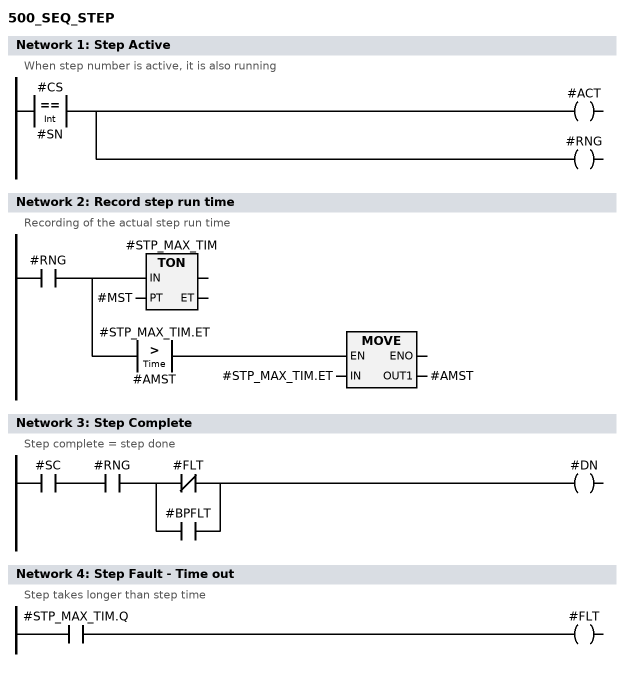
   RUNG wire#powerrail
      { S7_Templates := "SrcType := Int" } EQ_Contact(in1 := #CS, in2 := #SN)
      wire#w1
      Coil( #ACT )
   END_RUNG
   RUNG wire#w1
      Coil( #RNG )
   END_RUNG
   // the same network as SCL:
   #ACT := #CS = #SN;
   #RNG := #ACT;
END_REGION

REGION Network 2: Record step run time
   // Recording of the actual step run time
   #STP_MAX_TIM(IN := #RNG, PT := #MST);   // TON
   IF #RNG AND (#STP_MAX_TIM.ET > #AMST) THEN #AMST := #STP_MAX_TIM.ET; END_IF;
END_REGION

REGION Network 3: Step Complete
   // Step complete = step done
   RUNG wire#powerrail
      Contact( #SC )
      Contact( #RNG )
      wire#w1
      I_Contact( #FLT )
      wire#w2
      Coil( #DN )
   END_RUNG
   RUNG wire#w1
      Contact( #BPFLT )
   END_RUNG wire#w2
   // the same network as SCL:
   #DN := #SC AND #RNG AND (NOT #FLT OR #BPFLT);
END_REGION

REGION Network 4: Step Fault - Time out
   // Step takes longer than step time
   RUNG wire#powerrail
      Contact( #STP_MAX_TIM.Q )
      Coil( #FLT )
   END_RUNG
   // the same network as SCL:
   #FLT := #STP_MAX_TIM.Q;
END_REGION
END_FUNCTION_BLOCK

FUNCTION_BLOCK "501_VLV_CHK"   // FB501, LAD
TITLE = Valve Check
{ S7_Optimized_Access := 'TRUE' }
AUTHOR : JRS
VERSION : 0.1
// To check for the correct operation of a vlave
   VAR_INPUT
      DMND : Bool;   // Demand
      NO_TYPE : Bool;   // Valve type = open without demand
      NC_TYPE : Bool;   // Valve type = closed without demand
      MAX_MOV_TIM : Time := T#1s;   // Maximum movement time
      OPN_SNSR : Bool;   // Valve open confirmed
      CLS_SNSR : Bool;   // Valve closed confirmed
   END_VAR
   VAR_OUTPUT
      HELTHY : Bool;   // Valve is healthy
      FAULT : Bool;   // Valve is faulty
      CNFG_ERR : Bool;   // Configuration error
   END_VAR
   VAR
      IDLE_FLT : Bool;   // No demand fault
      DMND_FLT : Bool;   // Demand fault
      TRVL_TIME_FLT : Bool;   // Both sensors missing
      SNSR_FLT : Bool;   // Sensor conflicts
      TRVL_TIME : TON_TIME;   // Travel timer
   END_VAR
   // TRVL_TIME.PT := T#1s;
BEGIN

REGION Network 1: Idle Fault
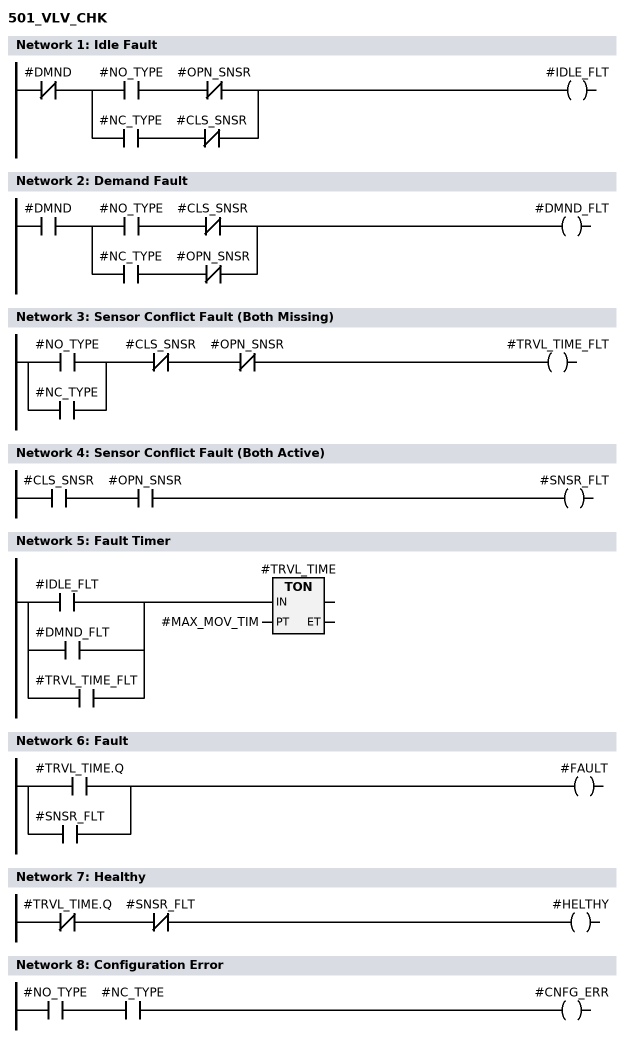
   RUNG wire#powerrail
      I_Contact( #DMND )
      wire#w1
      Contact( #NO_TYPE )
      I_Contact( #OPN_SNSR )
      wire#w2
      Coil( #IDLE_FLT )
   END_RUNG
   RUNG wire#w1
      Contact( #NC_TYPE )
      I_Contact( #CLS_SNSR )
   END_RUNG wire#w2
   // the same network as SCL:
   #IDLE_FLT := NOT #DMND AND ((#NO_TYPE AND NOT #OPN_SNSR) OR (#NC_TYPE AND NOT #CLS_SNSR));
END_REGION

REGION Network 2: Demand Fault
   RUNG wire#powerrail
      Contact( #DMND )
      wire#w1
      Contact( #NO_TYPE )
      I_Contact( #CLS_SNSR )
      wire#w2
      Coil( #DMND_FLT )
   END_RUNG
   RUNG wire#w1
      Contact( #NC_TYPE )
      I_Contact( #OPN_SNSR )
   END_RUNG wire#w2
   // the same network as SCL:
   #DMND_FLT := #DMND AND ((#NO_TYPE AND NOT #CLS_SNSR) OR (#NC_TYPE AND NOT #OPN_SNSR));
END_REGION

REGION Network 3: Sensor Conflict Fault (Both Missing)
   RUNG wire#powerrail
      Contact( #NO_TYPE )
      wire#w1
      I_Contact( #CLS_SNSR )
      I_Contact( #OPN_SNSR )
      Coil( #TRVL_TIME_FLT )
   END_RUNG
   RUNG wire#powerrail
      Contact( #NC_TYPE )
   END_RUNG wire#w1
   // the same network as SCL:
   #TRVL_TIME_FLT := (#NO_TYPE OR #NC_TYPE) AND NOT #CLS_SNSR AND NOT #OPN_SNSR;
END_REGION

REGION Network 4: Sensor Conflict Fault (Both Active)
   RUNG wire#powerrail
      Contact( #CLS_SNSR )
      Contact( #OPN_SNSR )
      Coil( #SNSR_FLT )
   END_RUNG
   // the same network as SCL:
   #SNSR_FLT := #CLS_SNSR AND #OPN_SNSR;
END_REGION

REGION Network 5: Fault Timer
   #TRVL_TIME(IN := #IDLE_FLT OR #DMND_FLT OR #TRVL_TIME_FLT, PT := #MAX_MOV_TIM);   // TON
END_REGION

REGION Network 6: Fault
   RUNG wire#powerrail
      Contact( #TRVL_TIME.Q )
      wire#w1
      Coil( #FAULT )
   END_RUNG
   RUNG wire#powerrail
      Contact( #SNSR_FLT )
   END_RUNG wire#w1
   // the same network as SCL:
   #FAULT := #TRVL_TIME.Q OR #SNSR_FLT;
END_REGION

REGION Network 7: Healthy
   RUNG wire#powerrail
      I_Contact( #TRVL_TIME.Q )
      I_Contact( #SNSR_FLT )
      Coil( #HELTHY )
   END_RUNG
   // the same network as SCL:
   #HELTHY := NOT #TRVL_TIME.Q AND NOT #SNSR_FLT;
END_REGION

REGION Network 8: Configuration Error
   RUNG wire#powerrail
      Contact( #NO_TYPE )
      Contact( #NC_TYPE )
      Coil( #CNFG_ERR )
   END_RUNG
   // the same network as SCL:
   #CNFG_ERR := #NO_TYPE AND #NC_TYPE;
END_REGION
END_FUNCTION_BLOCK

FUNCTION_BLOCK "502_ALM_ANALOG"   // FB502, LAD
{ S7_Optimized_Access := 'FALSE' }
VERSION : 0.1
   VAR_INPUT
      Value : Real;
      "Raw Value" : Int;
      Enable : Bool := true;
      "Enable Delay Time" : Time := T#10s;
      "High Value Release" : Bool := true;   // It is Releasing High Values from Enable restriction
      "SHORT CIRCUIT VALUE" : Real := 32000.0;
      "BROKEN WIRE VALUE" : Real := -32000.0;
      "VERY LOW LEVEL VALUE (LL)" : Real;
      "LOW LEVEL VALUE (L)" : Real;
      "HIGH LEVEL VALUE (H)" : Real;
      "VERY HIGH LEVEL VALUE (HH)" : Real;
      OFFSET : Real;
      "ALARM DELAY" : Time := T#1s;
      "Peak Value Reset" : Bool;
   END_VAR
   VAR_OUTPUT
      "ALARM HH" : Bool;
      "ALARM H" : Bool;
      "ALARM L" : Bool;
      "ALARM LL" : Bool;
      "ALARM READING" : Bool;
      "Peak Value" : Real;
      Alarm : Word;
      Alarm_INT : Int;
   END_VAR
   VAR
      TRUE : Bool;
      FALSE : Bool;
      Raw_value_int : Int;
      RET_VAL : Word;
      RAW_scaled_mA : Real;
      RAW_scaled_VALUE : Real;
      SCALED_OFFSETTED_VALUE : Real;
      Error_present : Bool;
      "Enable Internal" : Bool;
      "ALARM HH_interm" : Bool;
      "ALARM H_interm" : Bool;
      "ALARM L_interm" : Bool;
      "ALARM LL_interm" : Bool;
      "ALARM READING_interm" : Bool;
      "ALARM_HH delay" : TON_TIME;
      "ALARM_H delay" : TON_TIME;
      "ALARM_LL delay" : TON_TIME;
      "ALARM_L delay" : TON_TIME;
      "ALARM_READING delay" : TON_TIME;
      "ALARM READING TOF" : TOF_TIME;
      "HI HI TOF" : TOF_TIME;
      "HI TOF" : TOF_TIME;
      "LOE TOF" : TOF_TIME;
      "LOW TOF" : TOF_TIME;
      "LOW LOW TOF" : TOF_TIME;
      "Enable TON" : TON_TIME;
   END_VAR
   VAR_TEMP   // added for the SCL form of the ladder/FBD networks
      _w1 : Bool;
   END_VAR
BEGIN

REGION Network 1: True False
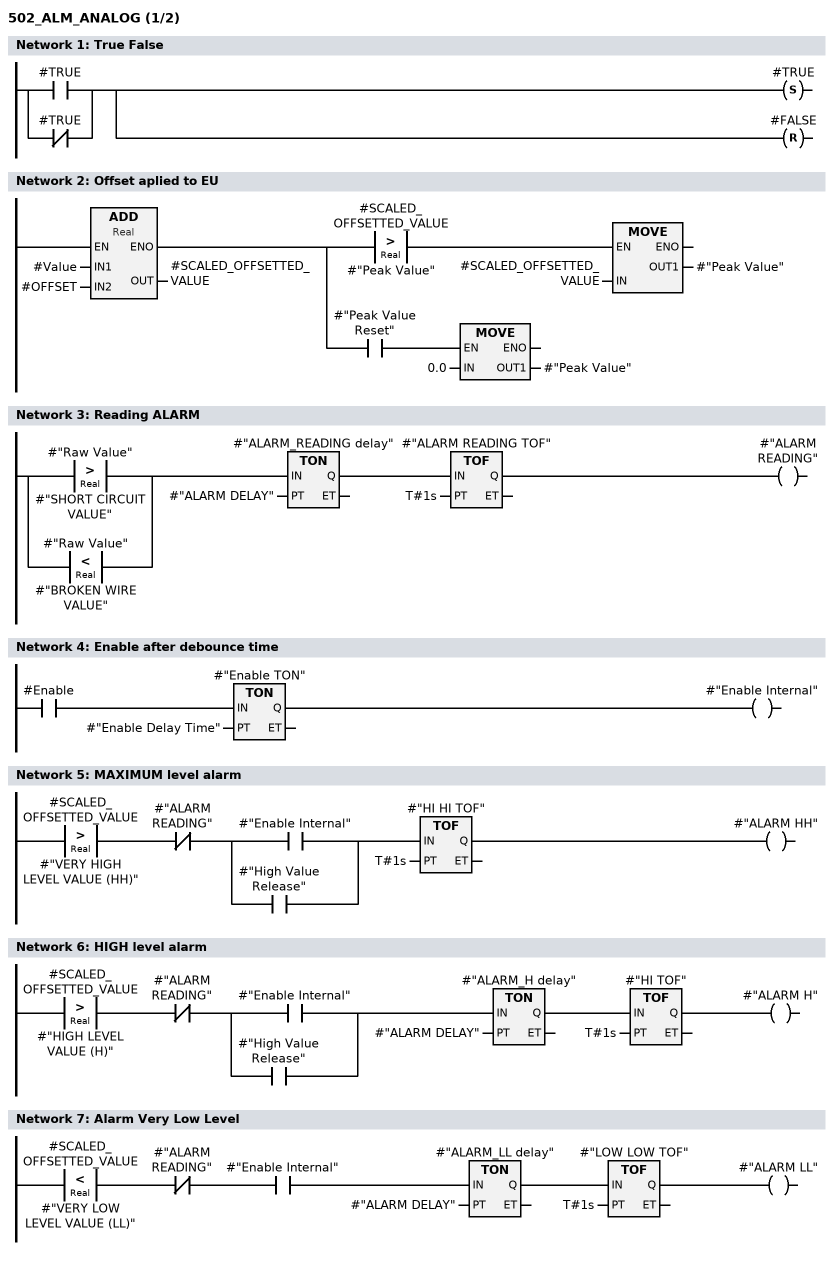
   RUNG wire#powerrail
      Contact( #TRUE )
      wire#w1
      S_Coil( #TRUE )
   END_RUNG
   RUNG wire#powerrail
      I_Contact( #TRUE )
   END_RUNG wire#w1
   RUNG wire#w1
      R_Coil( #FALSE )
   END_RUNG
   // the same network as SCL:
   #_w1 := #TRUE OR NOT #TRUE;
   IF #_w1 THEN
       #TRUE := TRUE;
       #FALSE := FALSE;
   END_IF;
END_REGION

REGION Network 2: Offset aplied to EU
   RUNG wire#powerrail
      { S7_Templates := "SrcType := Real"; S7_GenerateENO := "TRUE" } Add(in1 := #Value, in2 := #OFFSET, out => #SCALED_OFFSETTED_VALUE)
      wire#w1
      { S7_Templates := "SrcType := Real" } GT_Contact(in1 := #SCALED_OFFSETTED_VALUE, in2 := #"Peak Value")
      Move(in := #SCALED_OFFSETTED_VALUE, out1 => #"Peak Value")
   END_RUNG
   RUNG wire#w1
      Contact( #"Peak Value Reset" )
      Move(in := 0.0, out1 => #"Peak Value")
   END_RUNG
   // the same network as SCL:
   // ENO of a box is taken as its EN; it also drops when the box reports an error
   #SCALED_OFFSETTED_VALUE := #Value + #OFFSET;
   IF #SCALED_OFFSETTED_VALUE > #"Peak Value" THEN #"Peak Value" := #SCALED_OFFSETTED_VALUE; END_IF;
   IF #"Peak Value Reset" THEN #"Peak Value" := 0.0; END_IF;
END_REGION

REGION Network 3: Reading ALARM
   #"ALARM_READING delay"(IN := (#"Raw Value" > #"SHORT CIRCUIT VALUE") OR (#"Raw Value" < #"BROKEN WIRE VALUE"),   // TON
                          PT := #"ALARM DELAY");
   #"ALARM READING TOF"(IN := #"ALARM_READING delay".Q, PT := T#1s);   // TOF
   #"ALARM READING" := #"ALARM READING TOF".Q;
END_REGION

REGION Network 4: Enable after debounce time
   #"Enable TON"(IN := #Enable, PT := #"Enable Delay Time");   // TON
   #"Enable Internal" := #"Enable TON".Q;
END_REGION

REGION Network 5: MAXIMUM level alarm
   #"HI HI TOF"(IN := (#SCALED_OFFSETTED_VALUE > #"VERY HIGH LEVEL VALUE (HH)") AND NOT #"ALARM READING" AND (#"Enable Internal" OR #"High Value Release"),   // TOF
                PT := T#1s);
   #"ALARM HH" := #"HI HI TOF".Q;
END_REGION

REGION Network 6: HIGH level alarm
   #"ALARM_H delay"(IN := (#SCALED_OFFSETTED_VALUE > #"HIGH LEVEL VALUE (H)") AND NOT #"ALARM READING" AND (#"Enable Internal" OR #"High Value Release"),   // TON
                    PT := #"ALARM DELAY");
   #"HI TOF"(IN := #"ALARM_H delay".Q, PT := T#1s);   // TOF
   #"ALARM H" := #"HI TOF".Q;
END_REGION

REGION Network 7: Alarm Very Low Level
   #"ALARM_LL delay"(IN := (#SCALED_OFFSETTED_VALUE < #"VERY LOW LEVEL VALUE (LL)") AND NOT #"ALARM READING" AND #"Enable Internal",   // TON
                     PT := #"ALARM DELAY");
   #"LOW LOW TOF"(IN := #"ALARM_LL delay".Q, PT := T#1s);   // TOF
   #"ALARM LL" := #"LOW LOW TOF".Q;
END_REGION

REGION Network 8: Alarm Low Level
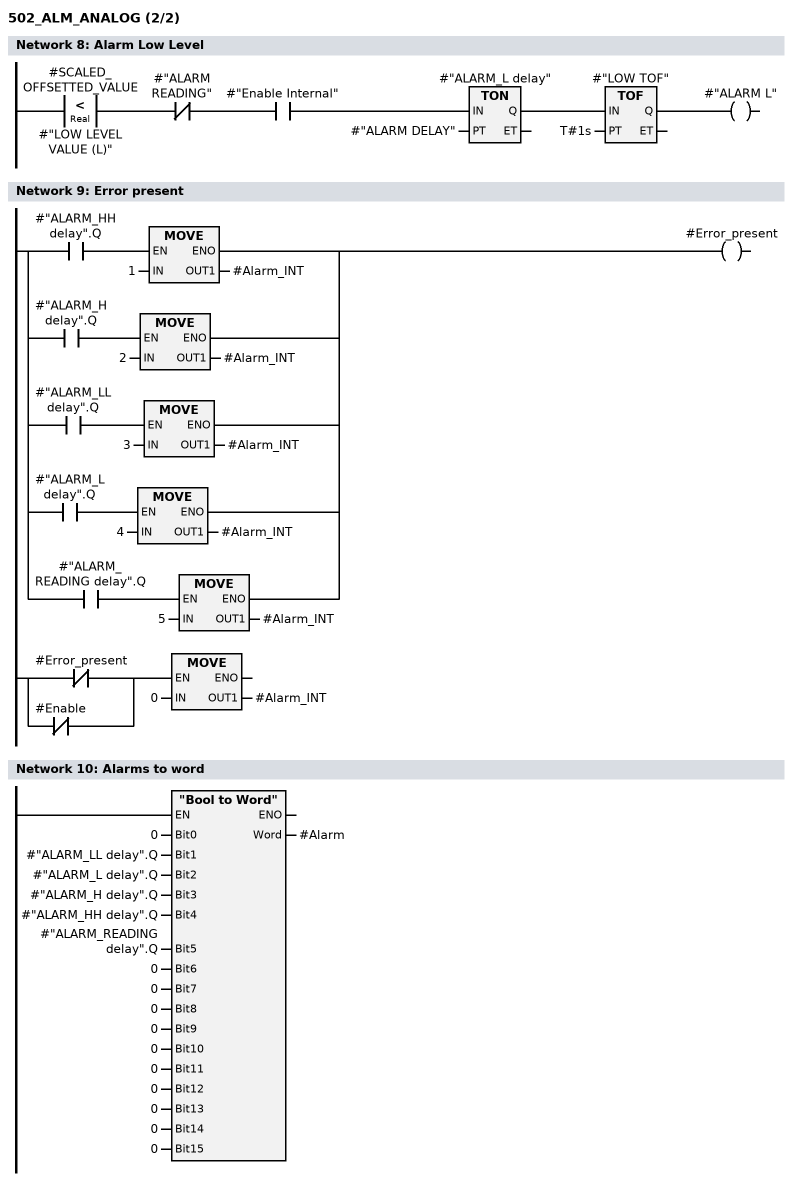
   #"ALARM_L delay"(IN := (#SCALED_OFFSETTED_VALUE < #"LOW LEVEL VALUE (L)") AND NOT #"ALARM READING" AND #"Enable Internal",   // TON
                    PT := #"ALARM DELAY");
   #"LOW TOF"(IN := #"ALARM_L delay".Q, PT := T#1s);   // TOF
   #"ALARM L" := #"LOW TOF".Q;
END_REGION

REGION Network 9: Error present
   RUNG wire#powerrail
      Contact( #"ALARM_HH delay".Q )
      { S7_GenerateENO := "TRUE" } Move(in := 1, out1 => #Alarm_INT)
      wire#w1
      Coil( #Error_present )
   END_RUNG
   RUNG wire#powerrail
      Contact( #"ALARM_H delay".Q )
      { S7_GenerateENO := "TRUE" } Move(in := 2, out1 => #Alarm_INT)
   END_RUNG wire#w1
   RUNG wire#powerrail
      Contact( #"ALARM_LL delay".Q )
      { S7_GenerateENO := "TRUE" } Move(in := 3, out1 => #Alarm_INT)
   END_RUNG wire#w1
   RUNG wire#powerrail
      Contact( #"ALARM_L delay".Q )
      { S7_GenerateENO := "TRUE" } Move(in := 4, out1 => #Alarm_INT)
   END_RUNG wire#w1
   RUNG wire#powerrail
      Contact( #"ALARM_READING delay".Q )
      { S7_GenerateENO := "TRUE" } Move(in := 5, out1 => #Alarm_INT)
   END_RUNG wire#w1
   RUNG wire#powerrail
      I_Contact( #Error_present )
      wire#w2
      Move(in := 0, out1 => #Alarm_INT)
   END_RUNG
   RUNG wire#powerrail
      I_Contact( #Enable )
   END_RUNG wire#w2
   // the same network as SCL:
   // ENO of a box is taken as its EN; it also drops when the box reports an error
   IF #"ALARM_HH delay".Q THEN #Alarm_INT := 1; END_IF;
   IF #"ALARM_H delay".Q THEN #Alarm_INT := 2; END_IF;
   IF #"ALARM_LL delay".Q THEN #Alarm_INT := 3; END_IF;
   IF #"ALARM_L delay".Q THEN #Alarm_INT := 4; END_IF;
   IF #"ALARM_READING delay".Q THEN #Alarm_INT := 5; END_IF;
   #Error_present := #"ALARM_HH delay".Q OR #"ALARM_H delay".Q OR #"ALARM_LL delay".Q OR #"ALARM_L delay".Q OR #"ALARM_READING delay".Q;
   IF NOT #Error_present OR NOT #Enable THEN #Alarm_INT := 0; END_IF;
END_REGION

REGION Network 10: Alarms to word
   RUNG wire#powerrail
      "Bool to Word"(Bit0 := 0, Bit1 := #"ALARM_LL delay".Q, Bit2 := #"ALARM_L delay".Q, Bit3 := #"ALARM_H delay".Q, Bit4 := #"ALARM_HH delay".Q, Bit5 := #"ALARM_READING delay".Q, Bit6 := 0, Bit7 := 0, Bit8 := 0, Bit9 := 0, Bit10 := 0, Bit11 := 0, Bit12 := 0, Bit13 := 0, Bit14 := 0, Bit15 := 0, "Word" => #Alarm)
   END_RUNG
   // the same network as SCL:
   "Bool to Word"(Bit0 := 0,
                  Bit1 := #"ALARM_LL delay".Q,
                  Bit2 := #"ALARM_L delay".Q,
                  Bit3 := #"ALARM_H delay".Q,
                  Bit4 := #"ALARM_HH delay".Q,
                  Bit5 := #"ALARM_READING delay".Q,
                  Bit6 := 0,
                  Bit7 := 0,
                  Bit8 := 0,
                  Bit9 := 0,
                  Bit10 := 0,
                  Bit11 := 0,
                  Bit12 := 0,
                  Bit13 := 0,
                  Bit14 := 0,
                  Bit15 := 0,
                  "Word" => #Alarm);
END_REGION
END_FUNCTION_BLOCK

FUNCTION_BLOCK "Alarm beacon handling"   // FB503, LAD
{ S7_Optimized_Access := 'TRUE' }
VERSION : 0.1
   VAR_INPUT
      Alarm : Bool;
      Warning : Bool;
      Latched : Bool;
      "Reset Alarm" : Bool;
      "Buzzer snooze" : Bool;
      "Beacon frequency" : Time;
      "Buzzer reset time" : Time;
   END_VAR
   VAR_OUTPUT
      "Alarm beacon" : Bool;
      "Warning beacon" : Bool;
      Buzzer : Bool;
      "Buzzer UnMute" : Bool;
   END_VAR
   VAR
      ON_Timer_0_Instance : TON_TIME;
      OFF_Timer_0_Instance : TON_TIME;
      Buzzer_Timer_0_Instance : TON_TIME;
      Alarm_interm : Bool;
      Warning_interm : Bool;
      "Reset Alarm Interm" : Bool;
      Aux1 : Bool;
      Aux2 : Bool;
      Aux3 : Bool;
      "Snooze Alarm" : Bool;
      "Snooze Warning" : Bool;
      "Alarm&Estop" : Bool;
   END_VAR
   VAR_TEMP   // added for the SCL form of the ladder/FBD networks
      _w1 : Bool;
      _w2 : Bool;
   END_VAR
BEGIN

REGION Network 1
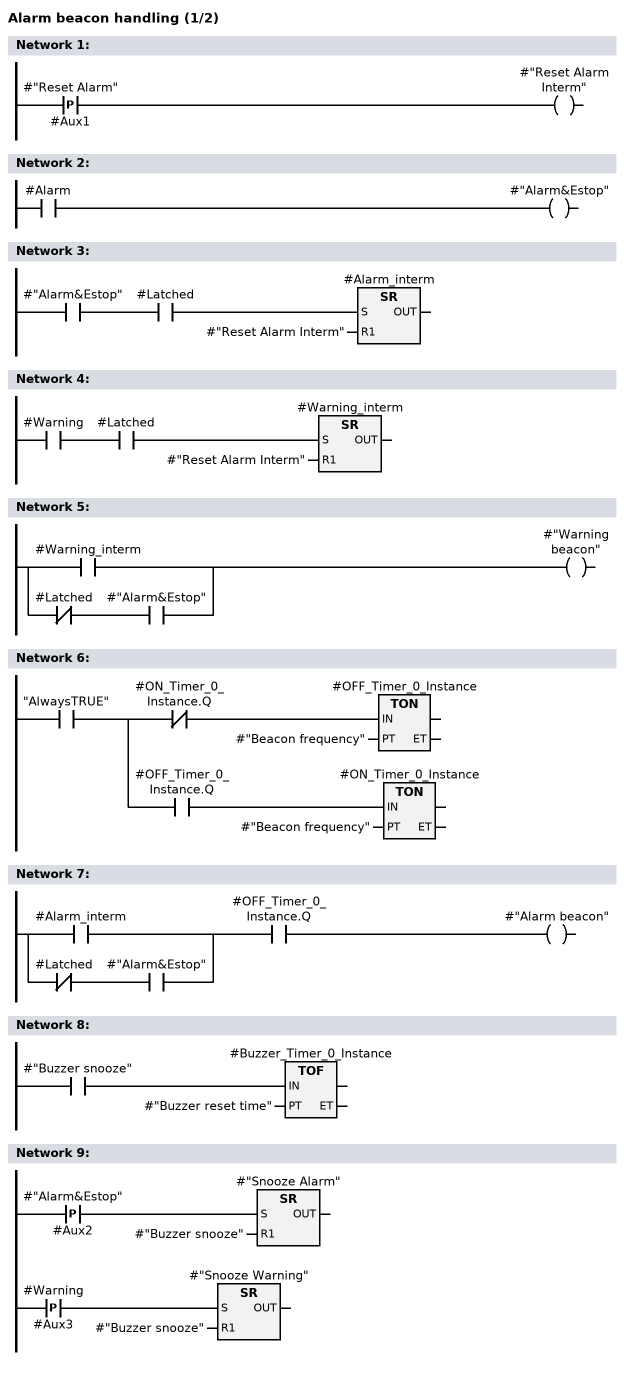
   RUNG wire#powerrail
      P_Contact(operand := #"Reset Alarm", bit := #Aux1)
      Coil( #"Reset Alarm Interm" )
   END_RUNG
   // the same network as SCL:
   #_w1 := #"Reset Alarm" AND NOT #Aux1;   // rising edge of #"Reset Alarm"
   #Aux1 := #"Reset Alarm";
   #"Reset Alarm Interm" := #_w1;
END_REGION

REGION Network 2
   RUNG wire#powerrail
      Contact( #Alarm )
      Coil( #"Alarm&Estop" )
   END_RUNG
   // the same network as SCL:
   #"Alarm&Estop" := #Alarm;
END_REGION

REGION Network 3
   RUNG wire#powerrail
      Contact( #"Alarm&Estop" )
      Contact( #Latched )
      S_SR(operand := #Alarm_interm, r1 := #"Reset Alarm Interm")
   END_RUNG
   // the same network as SCL:
   IF #"Alarm&Estop" AND #Latched THEN
       #Alarm_interm := TRUE;   // SR flip-flop
   END_IF;
   IF #"Reset Alarm Interm" THEN #Alarm_interm := FALSE; END_IF;
END_REGION

REGION Network 4
   RUNG wire#powerrail
      Contact( #Warning )
      Contact( #Latched )
      S_SR(operand := #Warning_interm, r1 := #"Reset Alarm Interm")
   END_RUNG
   // the same network as SCL:
   IF #Warning AND #Latched THEN
       #Warning_interm := TRUE;   // SR flip-flop
   END_IF;
   IF #"Reset Alarm Interm" THEN #Warning_interm := FALSE; END_IF;
END_REGION

REGION Network 5
   RUNG wire#powerrail
      Contact( #Warning_interm )
      wire#w1
      Coil( #"Warning beacon" )
   END_RUNG
   RUNG wire#powerrail
      I_Contact( #Latched )
      Contact( #"Alarm&Estop" )
   END_RUNG wire#w1
   // the same network as SCL:
   #"Warning beacon" := #Warning_interm OR (NOT #Latched AND #"Alarm&Estop");
END_REGION

REGION Network 6
   #OFF_Timer_0_Instance(IN := "AlwaysTRUE" AND NOT #ON_Timer_0_Instance.Q, PT := #"Beacon frequency");   // TON
   #ON_Timer_0_Instance(IN := "AlwaysTRUE" AND #OFF_Timer_0_Instance.Q, PT := #"Beacon frequency");   // TON
END_REGION

REGION Network 7
   RUNG wire#powerrail
      Contact( #Alarm_interm )
      wire#w1
      Contact( #OFF_Timer_0_Instance.Q )
      Coil( #"Alarm beacon" )
   END_RUNG
   RUNG wire#powerrail
      I_Contact( #Latched )
      Contact( #"Alarm&Estop" )
   END_RUNG wire#w1
   // the same network as SCL:
   #"Alarm beacon" := (#Alarm_interm OR (NOT #Latched AND #"Alarm&Estop")) AND #OFF_Timer_0_Instance.Q;
END_REGION

REGION Network 8
   #Buzzer_Timer_0_Instance(IN := #"Buzzer snooze", PT := #"Buzzer reset time");   // TOF
END_REGION

REGION Network 9
   RUNG wire#powerrail
      P_Contact(operand := #"Alarm&Estop", bit := #Aux2)
      S_SR(operand := #"Snooze Alarm", r1 := #"Buzzer snooze")
   END_RUNG
   RUNG wire#powerrail
      P_Contact(operand := #Warning, bit := #Aux3)
      S_SR(operand := #"Snooze Warning", r1 := #"Buzzer snooze")
   END_RUNG
   // the same network as SCL:
   #_w1 := #"Alarm&Estop" AND NOT #Aux2;   // rising edge of #"Alarm&Estop"
   #Aux2 := #"Alarm&Estop";
   IF #_w1 THEN
       #"Snooze Alarm" := TRUE;   // SR flip-flop
   END_IF;
   IF #"Buzzer snooze" THEN #"Snooze Alarm" := FALSE; END_IF;
   #_w2 := #Warning AND NOT #Aux3;   // rising edge of #Warning
   #Aux3 := #Warning;
   IF #_w2 THEN
       #"Snooze Warning" := TRUE;   // SR flip-flop
   END_IF;
   IF #"Buzzer snooze" THEN #"Snooze Warning" := FALSE; END_IF;
END_REGION

REGION Network 10
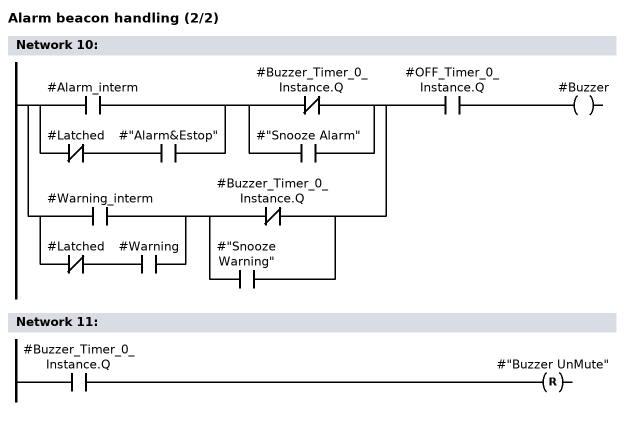
   RUNG wire#powerrail
      Contact( #Alarm_interm )
      wire#w1
      I_Contact( #Buzzer_Timer_0_Instance.Q )
      wire#w2
      Contact( #OFF_Timer_0_Instance.Q )
      Coil( #Buzzer )
   END_RUNG
   RUNG wire#powerrail
      I_Contact( #Latched )
      Contact( #"Alarm&Estop" )
   END_RUNG wire#w1
   RUNG wire#w1
      Contact( #"Snooze Alarm" )
   END_RUNG wire#w2
   RUNG wire#powerrail
      Contact( #Warning_interm )
      wire#w3
      I_Contact( #Buzzer_Timer_0_Instance.Q )
   END_RUNG wire#w2
   RUNG wire#powerrail
      I_Contact( #Latched )
      Contact( #Warning )
   END_RUNG wire#w3
   RUNG wire#w3
      Contact( #"Snooze Warning" )
   END_RUNG wire#w2
   // the same network as SCL:
   #Buzzer := (((#Alarm_interm OR (NOT #Latched AND #"Alarm&Estop")) AND (NOT #Buzzer_Timer_0_Instance.Q OR #"Snooze Alarm")) OR ((#Warning_interm OR (NOT #Latched AND #Warning)) AND (NOT #Buzzer_Timer_0_Instance.Q OR #"Snooze Warning"))) AND #OFF_Timer_0_Instance.Q;
END_REGION

REGION Network 11
   RUNG wire#powerrail
      Contact( #Buzzer_Timer_0_Instance.Q )
      R_Coil( #"Buzzer UnMute" )
   END_RUNG
   // the same network as SCL:
   IF #Buzzer_Timer_0_Instance.Q THEN #"Buzzer UnMute" := FALSE; END_IF;
END_REGION
END_FUNCTION_BLOCK

FUNCTION_BLOCK "64_Functioning Hours"   // FB506, LAD
{ S7_Optimized_Access := 'TRUE' }
VERSION : 0.1
   VAR_INPUT
      Started : Bool;
      Reset : Bool;
      "Service Time Days" : Int;
      "Service Time Hours" : Int;
   END_VAR
   VAR_OUTPUT
      Seconds : Int;
      Minutes : Int;
      Hours : Int;
      Days : Int;
      "Second beat_bit" : Bool;
      "Service Time bit" : Bool;
      "Hours to Service" : Int;
      "Hours Total" : Int;
      "Hours Functioning_Out" : Int;
   END_VAR
   VAR
      "Second beat" : TON_TIME;
      "Second Reset" : TON_TIME;
   END_VAR
   VAR RETAIN
      "Seconds burn" : CTU_INT;
      "Minutes burn" : CTU_INT;
      "Hours burn" : CTU_INT;
      "Days burn" : CTU_INT;
      Aux : Struct
         Aux_1 : Bool;
         Aux_2 : Bool;
         Aux_3 : Bool;
         Aux_4 : Bool;
         Aux_Puls : Bool;
         Aux_PulsN : Bool;
         Aux_HoursFunctioning : Int;
         "Aux_Total Hours" : Int;
      END_STRUCT;
   END_VAR
   VAR
      "Hours Functioning" : Int;
   END_VAR
   VAR_TEMP   // added for the SCL form of the ladder/FBD networks
      _w1 : Bool;
      _w2 : Bool;
      _w3 : Bool;
   END_VAR
BEGIN

REGION Network 1
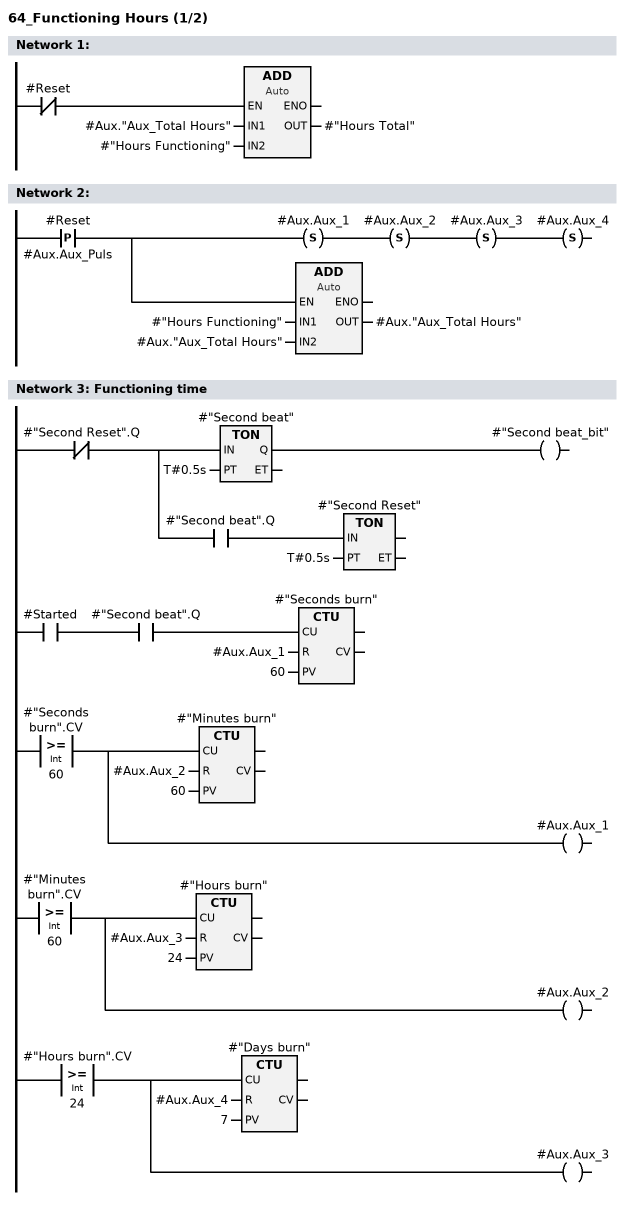
   RUNG wire#powerrail
      I_Contact( #Reset )
      Add(in1 := #Aux."Aux_Total Hours", in2 := #"Hours Functioning", out => #"Hours Total")
   END_RUNG
   // the same network as SCL:
   IF NOT #Reset THEN #"Hours Total" := #Aux."Aux_Total Hours" + #"Hours Functioning"; END_IF;
END_REGION

REGION Network 2
   RUNG wire#powerrail
      P_Contact(operand := #Reset, bit := #Aux.Aux_Puls)
      wire#w1
      S_Coil( #Aux.Aux_1 )
      S_Coil( #Aux.Aux_2 )
      S_Coil( #Aux.Aux_3 )
      S_Coil( #Aux.Aux_4 )
   END_RUNG
   RUNG wire#w1
      Add(in1 := #"Hours Functioning", in2 := #Aux."Aux_Total Hours", out => #Aux."Aux_Total Hours")
   END_RUNG
   // the same network as SCL:
   #_w1 := #Reset AND NOT #Aux.Aux_Puls;   // rising edge of #Reset
   #Aux.Aux_Puls := #Reset;
   IF #_w1 THEN
       #Aux.Aux_1 := TRUE;
       #Aux.Aux_2 := TRUE;
       #Aux.Aux_3 := TRUE;
       #Aux.Aux_4 := TRUE;
       #Aux."Aux_Total Hours" := #"Hours Functioning" + #Aux."Aux_Total Hours";
   END_IF;
END_REGION

REGION Network 3: Functioning time
   #"Second beat"(IN := NOT #"Second Reset".Q, PT := T#0.5s);   // TON
   #"Second beat_bit" := #"Second beat".Q;
   #"Second Reset"(IN := NOT #"Second Reset".Q AND #"Second beat".Q, PT := T#0.5s);   // TON
   #"Seconds burn"(CU := #Started AND #"Second beat".Q, R := #Aux.Aux_1, PV := 60);   // CTU
   #_w1 := #"Seconds burn".CV >= 60;
   #"Minutes burn"(CU := #_w1, R := #Aux.Aux_2, PV := 60);   // CTU
   #Aux.Aux_1 := #_w1;
   #_w2 := #"Minutes burn".CV >= 60;
   #"Hours burn"(CU := #_w2, R := #Aux.Aux_3, PV := 24);   // CTU
   #Aux.Aux_2 := #_w2;
   #_w3 := #"Hours burn".CV >= 24;
   #"Days burn"(CU := #_w3, R := #Aux.Aux_4, PV := 7);   // CTU
   #Aux.Aux_3 := #_w3;
END_REGION

REGION Network 4